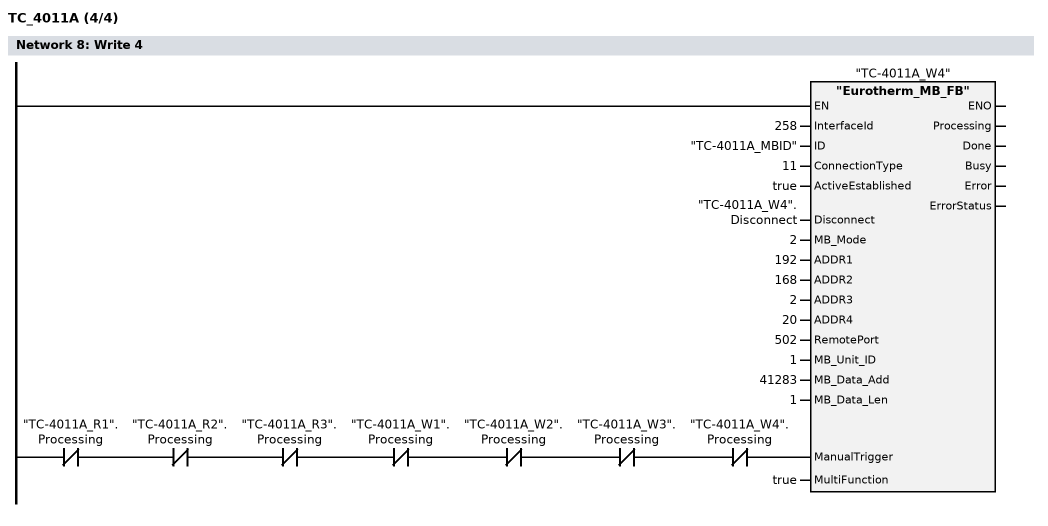
   RUNG wire#powerrail
      "TC-4011A_W4"(ManualTrigger := wire#w1, InterfaceId := 258, ID := "TC-4011A_MBID", ConnectionType := 11, ActiveEstablished := true, Disconnect := "TC-4011A_W4".Disconnect, MB_Mode := 2, ADDR1 := 192, ADDR2 := 168, ADDR3 := 2, ADDR4 := 20, RemotePort := 502, MB_Unit_ID := 1, MB_Data_Add := 41283, MB_Data_Len := 1, MultiFunction := true, Processing =>, Done =>, Busy =>, Error =>, ErrorStatus =>)
   END_RUNG
   RUNG wire#powerrail
      I_Contact( "TC-4011A_R1".Processing )
      I_Contact( "TC-4011A_R2".Processing )
      I_Contact( "TC-4011A_R3".Processing )
      I_Contact( "TC-4011A_W1".Processing )
      I_Contact( "TC-4011A_W2".Processing )
      I_Contact( "TC-4011A_W3".Processing )
      I_Contact( "TC-4011A_W4".Processing )
   END_RUNG wire#w1
   // the same network as SCL:
   "TC-4011A_W4"(InterfaceId := 258,   // "Eurotherm_MB_FB"
                 ID := "TC-4011A_MBID",
                 ConnectionType := 11,
                 ActiveEstablished := true,
                 Disconnect := "TC-4011A_W4".Disconnect,
                 MB_Mode := 2,
                 ADDR1 := 192,
                 ADDR2 := 168,
                 ADDR3 := 2,
                 ADDR4 := 20,
                 RemotePort := 502,
                 MB_Unit_ID := 1,
                 MB_Data_Add := 41283,
                 MB_Data_Len := 1,
                 ManualTrigger := NOT "TC-4011A_R1".Processing AND NOT "TC-4011A_R2".Processing AND NOT "TC-4011A_R3".Processing AND NOT "TC-4011A_W1".Processing AND NOT "TC-4011A_W2".Processing AND NOT "TC-4011A_W3".Processing AND NOT "TC-4011A_W4".Processing,
                 MultiFunction := true);
END_REGION
END_FUNCTION

// folder: Outside Comms/ModBus Comms/EurothermControllers/TC-4011B

FUNCTION "TC_4011B" : Void   // FC32, LAD
{ S7_Optimized_Access := 'TRUE' }
VERSION : 0.1
BEGIN

REGION Network 2: Read Data 1
   // R1=30001
   // R2=31280
   // R3=30023
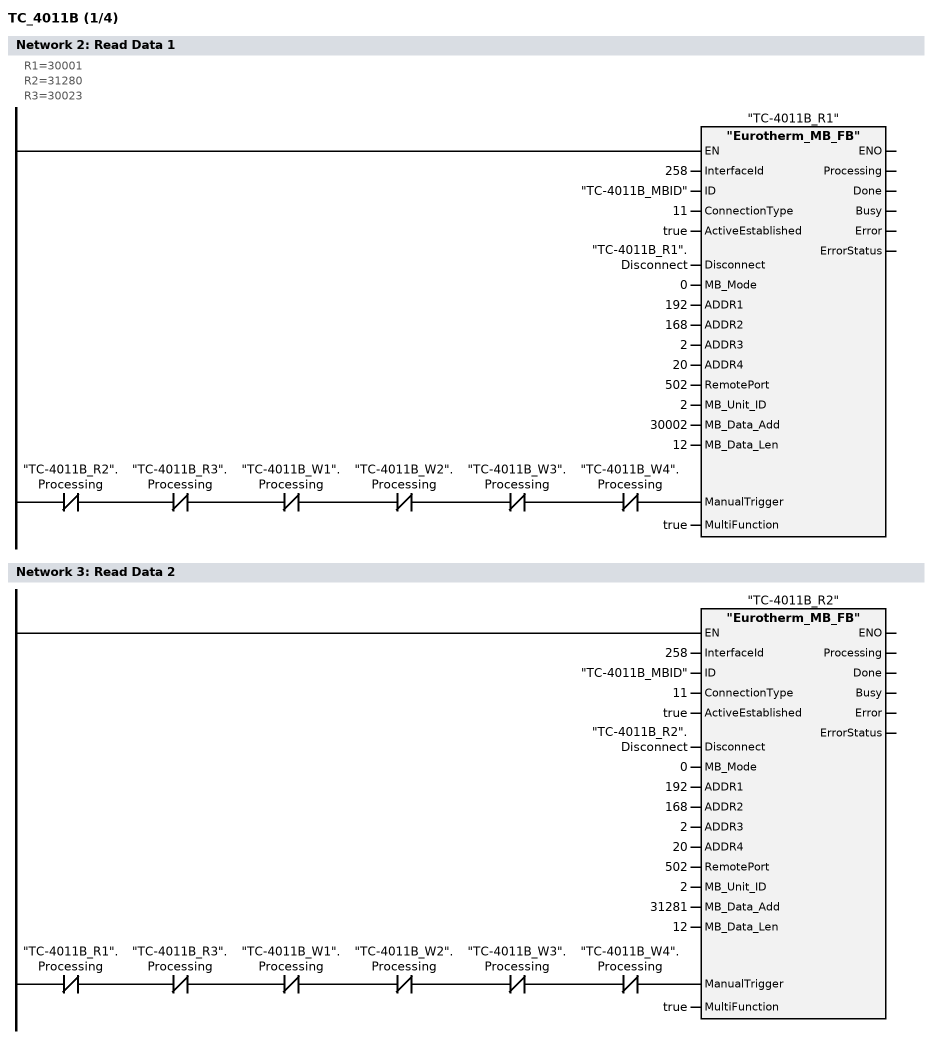
   RUNG wire#powerrail
      "TC-4011B_R1"(ManualTrigger := wire#w1, InterfaceId := 258, ID := "TC-4011B_MBID", ConnectionType := 11, ActiveEstablished := true, Disconnect := "TC-4011B_R1".Disconnect, MB_Mode := 0, ADDR1 := 192, ADDR2 := 168, ADDR3 := 2, ADDR4 := 20, RemotePort := 502, MB_Unit_ID := 2, MB_Data_Add := 30002, MB_Data_Len := 12, MultiFunction := true, Processing =>, Done =>, Busy =>, Error =>, ErrorStatus =>)
   END_RUNG
   RUNG wire#powerrail
      I_Contact( "TC-4011B_R2".Processing )
      I_Contact( "TC-4011B_R3".Processing )
      I_Contact( "TC-4011B_W1".Processing )
      I_Contact( "TC-4011B_W2".Processing )
      I_Contact( "TC-4011B_W3".Processing )
      I_Contact( "TC-4011B_W4".Processing )
   END_RUNG wire#w1
   // the same network as SCL:
   "TC-4011B_R1"(InterfaceId := 258,   // "Eurotherm_MB_FB"
                 ID := "TC-4011B_MBID",
                 ConnectionType := 11,
                 ActiveEstablished := true,
                 Disconnect := "TC-4011B_R1".Disconnect,
                 MB_Mode := 0,
                 ADDR1 := 192,
                 ADDR2 := 168,
                 ADDR3 := 2,
                 ADDR4 := 20,
                 RemotePort := 502,
                 MB_Unit_ID := 2,
                 MB_Data_Add := 30002,
                 MB_Data_Len := 12,
                 ManualTrigger := NOT "TC-4011B_R2".Processing AND NOT "TC-4011B_R3".Processing AND NOT "TC-4011B_W1".Processing AND NOT "TC-4011B_W2".Processing AND NOT "TC-4011B_W3".Processing AND NOT "TC-4011B_W4".Processing,
                 MultiFunction := true);
END_REGION

REGION Network 3: Read Data 2
   RUNG wire#powerrail
      "TC-4011B_R2"(ManualTrigger := wire#w1, InterfaceId := 258, ID := "TC-4011B_MBID", ConnectionType := 11, ActiveEstablished := true, Disconnect := "TC-4011B_R2".Disconnect, MB_Mode := 0, ADDR1 := 192, ADDR2 := 168, ADDR3 := 2, ADDR4 := 20, RemotePort := 502, MB_Unit_ID := 2, MB_Data_Add := 31281, MB_Data_Len := 12, MultiFunction := true, Processing =>, Done =>, Busy =>, Error =>, ErrorStatus =>)
   END_RUNG
   RUNG wire#powerrail
      I_Contact( "TC-4011B_R1".Processing )
      I_Contact( "TC-4011B_R3".Processing )
      I_Contact( "TC-4011B_W1".Processing )
      I_Contact( "TC-4011B_W2".Processing )
      I_Contact( "TC-4011B_W3".Processing )
      I_Contact( "TC-4011B_W4".Processing )
   END_RUNG wire#w1
   // the same network as SCL:
   "TC-4011B_R2"(InterfaceId := 258,   // "Eurotherm_MB_FB"
                 ID := "TC-4011B_MBID",
                 ConnectionType := 11,
                 ActiveEstablished := true,
                 Disconnect := "TC-4011B_R2".Disconnect,
                 MB_Mode := 0,
                 ADDR1 := 192,
                 ADDR2 := 168,
                 ADDR3 := 2,
                 ADDR4 := 20,
                 RemotePort := 502,
                 MB_Unit_ID := 2,
                 MB_Data_Add := 31281,
                 MB_Data_Len := 12,
                 ManualTrigger := NOT "TC-4011B_R1".Processing AND NOT "TC-4011B_R3".Processing AND NOT "TC-4011B_W1".Processing AND NOT "TC-4011B_W2".Processing AND NOT "TC-4011B_W3".Processing AND NOT "TC-4011B_W4".Processing,
                 MultiFunction := true);
END_REGION

REGION Network 4: Read Data 3
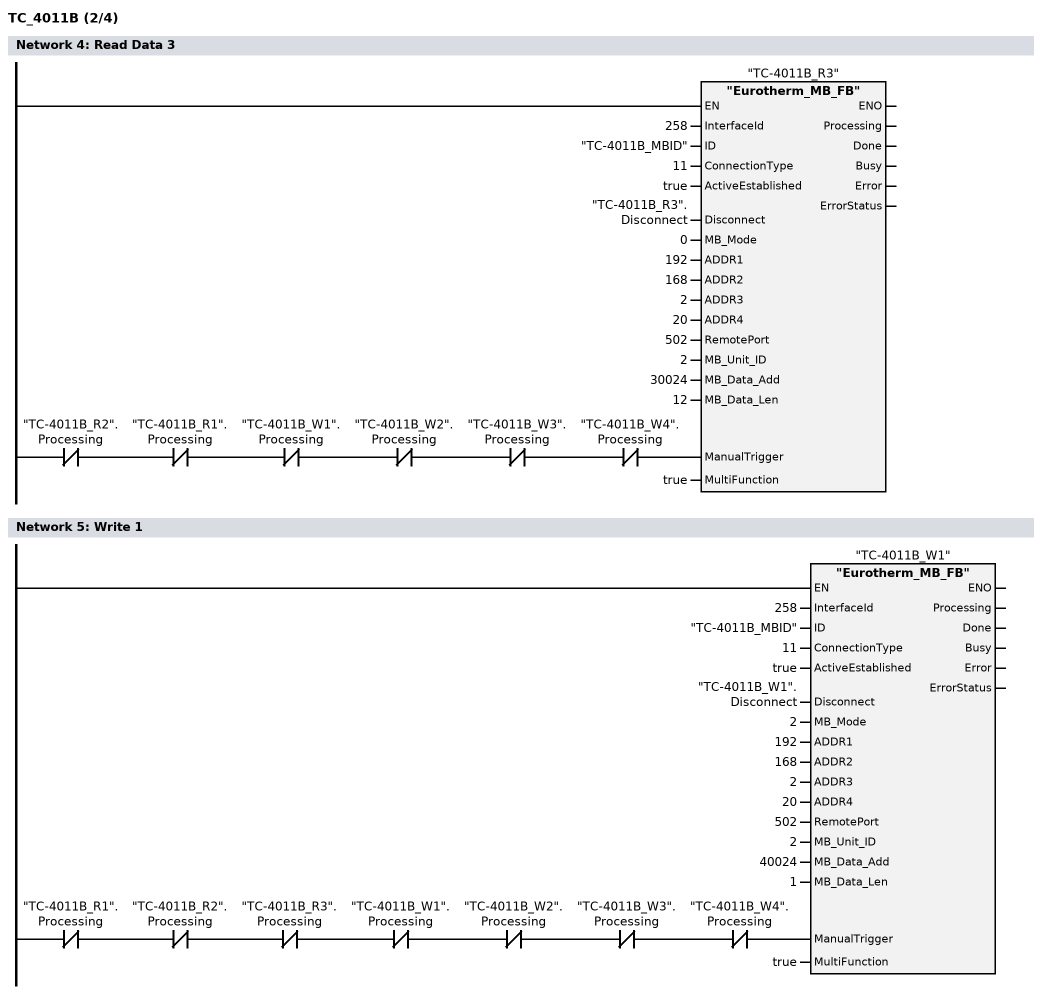
   RUNG wire#powerrail
      "TC-4011B_R3"(ManualTrigger := wire#w1, InterfaceId := 258, ID := "TC-4011B_MBID", ConnectionType := 11, ActiveEstablished := true, Disconnect := "TC-4011B_R3".Disconnect, MB_Mode := 0, ADDR1 := 192, ADDR2 := 168, ADDR3 := 2, ADDR4 := 20, RemotePort := 502, MB_Unit_ID := 2, MB_Data_Add := 30024, MB_Data_Len := 12, MultiFunction := true, Processing =>, Done =>, Busy =>, Error =>, ErrorStatus =>)
   END_RUNG
   RUNG wire#powerrail
      I_Contact( "TC-4011B_R2".Processing )
      I_Contact( "TC-4011B_R1".Processing )
      I_Contact( "TC-4011B_W1".Processing )
      I_Contact( "TC-4011B_W2".Processing )
      I_Contact( "TC-4011B_W3".Processing )
      I_Contact( "TC-4011B_W4".Processing )
   END_RUNG wire#w1
   // the same network as SCL:
   "TC-4011B_R3"(InterfaceId := 258,   // "Eurotherm_MB_FB"
                 ID := "TC-4011B_MBID",
                 ConnectionType := 11,
                 ActiveEstablished := true,
                 Disconnect := "TC-4011B_R3".Disconnect,
                 MB_Mode := 0,
                 ADDR1 := 192,
                 ADDR2 := 168,
                 ADDR3 := 2,
                 ADDR4 := 20,
                 RemotePort := 502,
                 MB_Unit_ID := 2,
                 MB_Data_Add := 30024,
                 MB_Data_Len := 12,
                 ManualTrigger := NOT "TC-4011B_R2".Processing AND NOT "TC-4011B_R1".Processing AND NOT "TC-4011B_W1".Processing AND NOT "TC-4011B_W2".Processing AND NOT "TC-4011B_W3".Processing AND NOT "TC-4011B_W4".Processing,
                 MultiFunction := true);
END_REGION

REGION Network 5: Write 1
   RUNG wire#powerrail
      "TC-4011B_W1"(ManualTrigger := wire#w1, InterfaceId := 258, ID := "TC-4011B_MBID", ConnectionType := 11, ActiveEstablished := true, Disconnect := "TC-4011B_W1".Disconnect, MB_Mode := 2, ADDR1 := 192, ADDR2 := 168, ADDR3 := 2, ADDR4 := 20, RemotePort := 502, MB_Unit_ID := 2, MB_Data_Add := 40024, MB_Data_Len := 1, MultiFunction := true, Processing =>, Done =>, Busy =>, Error =>, ErrorStatus =>)
   END_RUNG
   RUNG wire#powerrail
      I_Contact( "TC-4011B_R1".Processing )
      I_Contact( "TC-4011B_R2".Processing )
      I_Contact( "TC-4011B_R3".Processing )
      I_Contact( "TC-4011B_W1".Processing )
      I_Contact( "TC-4011B_W2".Processing )
      I_Contact( "TC-4011B_W3".Processing )
      I_Contact( "TC-4011B_W4".Processing )
   END_RUNG wire#w1
   // the same network as SCL:
   "TC-4011B_W1"(InterfaceId := 258,   // "Eurotherm_MB_FB"
                 ID := "TC-4011B_MBID",
                 ConnectionType := 11,
                 ActiveEstablished := true,
                 Disconnect := "TC-4011B_W1".Disconnect,
                 MB_Mode := 2,
                 ADDR1 := 192,
                 ADDR2 := 168,
                 ADDR3 := 2,
                 ADDR4 := 20,
                 RemotePort := 502,
                 MB_Unit_ID := 2,
                 MB_Data_Add := 40024,
                 MB_Data_Len := 1,
                 ManualTrigger := NOT "TC-4011B_R1".Processing AND NOT "TC-4011B_R2".Processing AND NOT "TC-4011B_R3".Processing AND NOT "TC-4011B_W1".Processing AND NOT "TC-4011B_W2".Processing AND NOT "TC-4011B_W3".Processing AND NOT "TC-4011B_W4".Processing,
                 MultiFunction := true);
END_REGION

REGION Network 6: Write 2
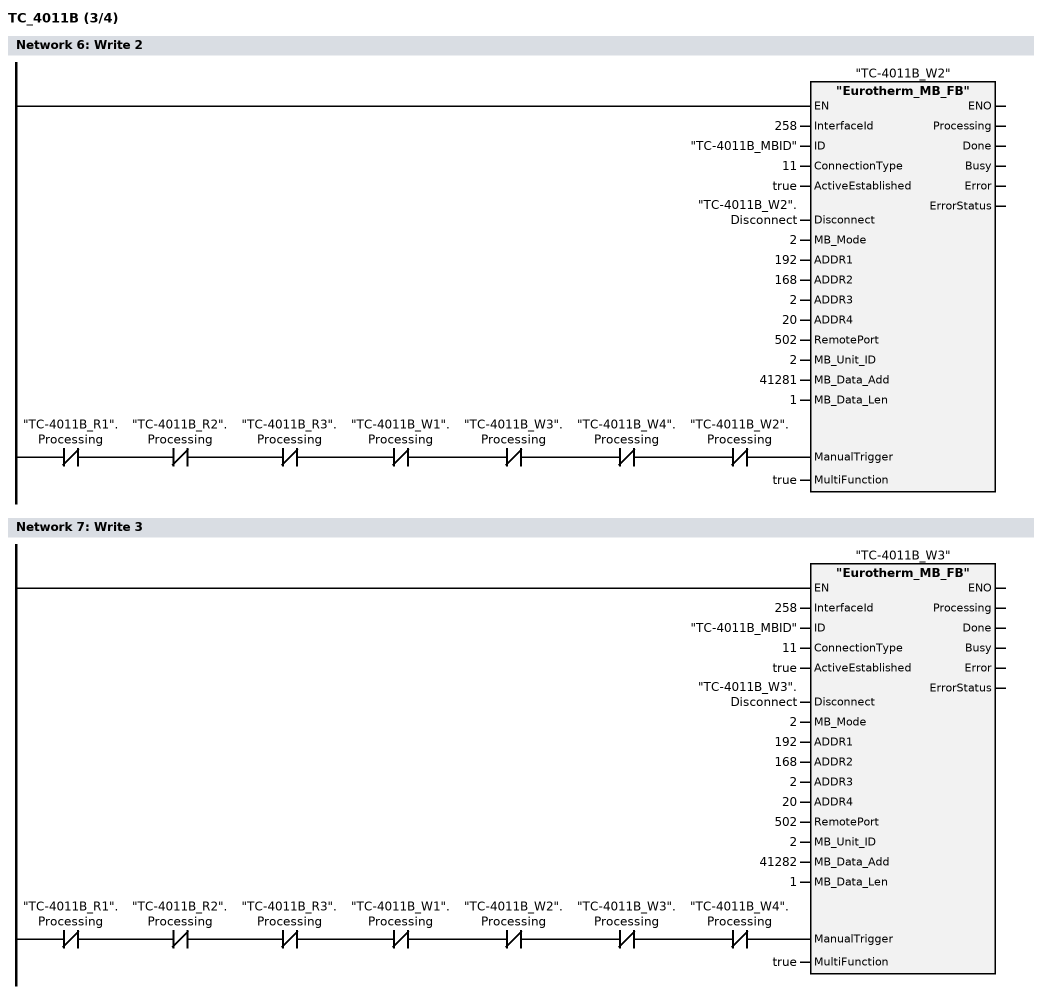
   RUNG wire#powerrail
      "TC-4011B_W2"(ManualTrigger := wire#w1, InterfaceId := 258, ID := "TC-4011B_MBID", ConnectionType := 11, ActiveEstablished := true, Disconnect := "TC-4011B_W2".Disconnect, MB_Mode := 2, ADDR1 := 192, ADDR2 := 168, ADDR3 := 2, ADDR4 := 20, RemotePort := 502, MB_Unit_ID := 2, MB_Data_Add := 41281, MB_Data_Len := 1, MultiFunction := true, Processing =>, Done =>, Busy =>, Error =>, ErrorStatus =>)
   END_RUNG
   RUNG wire#powerrail
      I_Contact( "TC-4011B_R1".Processing )
      I_Contact( "TC-4011B_R2".Processing )
      I_Contact( "TC-4011B_R3".Processing )
      I_Contact( "TC-4011B_W1".Processing )
      I_Contact( "TC-4011B_W3".Processing )
      I_Contact( "TC-4011B_W4".Processing )
      I_Contact( "TC-4011B_W2".Processing )
   END_RUNG wire#w1
   // the same network as SCL:
   "TC-4011B_W2"(InterfaceId := 258,   // "Eurotherm_MB_FB"
                 ID := "TC-4011B_MBID",
                 ConnectionType := 11,
                 ActiveEstablished := true,
                 Disconnect := "TC-4011B_W2".Disconnect,
                 MB_Mode := 2,
                 ADDR1 := 192,
                 ADDR2 := 168,
                 ADDR3 := 2,
                 ADDR4 := 20,
                 RemotePort := 502,
                 MB_Unit_ID := 2,
                 MB_Data_Add := 41281,
                 MB_Data_Len := 1,
                 ManualTrigger := NOT "TC-4011B_R1".Processing AND NOT "TC-4011B_R2".Processing AND NOT "TC-4011B_R3".Processing AND NOT "TC-4011B_W1".Processing AND NOT "TC-4011B_W3".Processing AND NOT "TC-4011B_W4".Processing AND NOT "TC-4011B_W2".Processing,
                 MultiFunction := true);
END_REGION

REGION Network 7: Write 3
   RUNG wire#powerrail
      "TC-4011B_W3"(ManualTrigger := wire#w1, InterfaceId := 258, ID := "TC-4011B_MBID", ConnectionType := 11, ActiveEstablished := true, Disconnect := "TC-4011B_W3".Disconnect, MB_Mode := 2, ADDR1 := 192, ADDR2 := 168, ADDR3 := 2, ADDR4 := 20, RemotePort := 502, MB_Unit_ID := 2, MB_Data_Add := 41282, MB_Data_Len := 1, MultiFunction := true, Processing =>, Done =>, Busy =>, Error =>, ErrorStatus =>)
   END_RUNG
   RUNG wire#powerrail
      I_Contact( "TC-4011B_R1".Processing )
      I_Contact( "TC-4011B_R2".Processing )
      I_Contact( "TC-4011B_R3".Processing )
      I_Contact( "TC-4011B_W1".Processing )
      I_Contact( "TC-4011B_W2".Processing )
      I_Contact( "TC-4011B_W3".Processing )
      I_Contact( "TC-4011B_W4".Processing )
   END_RUNG wire#w1
   // the same network as SCL:
   "TC-4011B_W3"(InterfaceId := 258,   // "Eurotherm_MB_FB"
                 ID := "TC-4011B_MBID",
                 ConnectionType := 11,
                 ActiveEstablished := true,
                 Disconnect := "TC-4011B_W3".Disconnect,
                 MB_Mode := 2,
                 ADDR1 := 192,
                 ADDR2 := 168,
                 ADDR3 := 2,
                 ADDR4 := 20,
                 RemotePort := 502,
                 MB_Unit_ID := 2,
                 MB_Data_Add := 41282,
                 MB_Data_Len := 1,
                 ManualTrigger := NOT "TC-4011B_R1".Processing AND NOT "TC-4011B_R2".Processing AND NOT "TC-4011B_R3".Processing AND NOT "TC-4011B_W1".Processing AND NOT "TC-4011B_W2".Processing AND NOT "TC-4011B_W3".Processing AND NOT "TC-4011B_W4".Processing,
                 MultiFunction := true);
END_REGION

REGION Network 8: Write 4
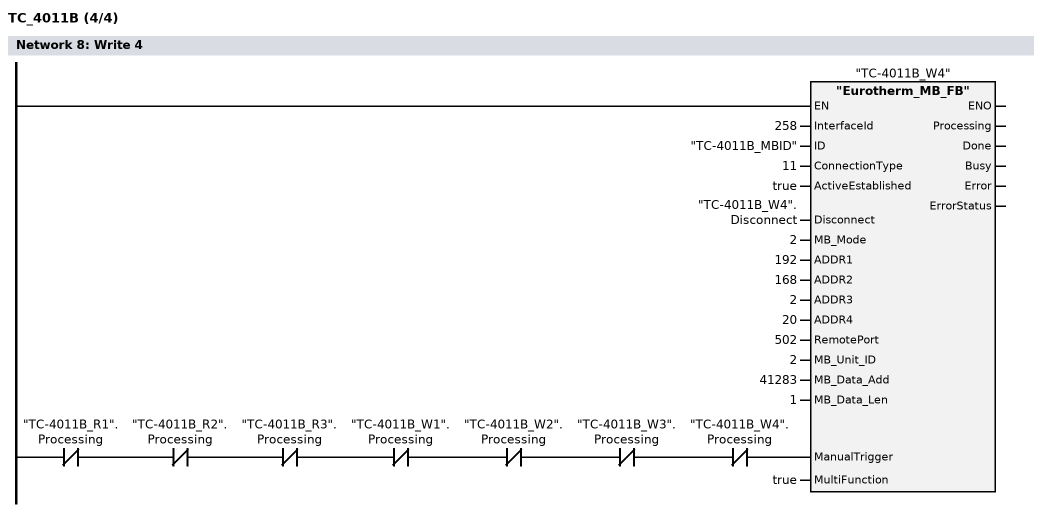
   RUNG wire#powerrail
      "TC-4011B_W4"(ManualTrigger := wire#w1, InterfaceId := 258, ID := "TC-4011B_MBID", ConnectionType := 11, ActiveEstablished := true, Disconnect := "TC-4011B_W4".Disconnect, MB_Mode := 2, ADDR1 := 192, ADDR2 := 168, ADDR3 := 2, ADDR4 := 20, RemotePort := 502, MB_Unit_ID := 2, MB_Data_Add := 41283, MB_Data_Len := 1, MultiFunction := true, Processing =>, Done =>, Busy =>, Error =>, ErrorStatus =>)
   END_RUNG
   RUNG wire#powerrail
      I_Contact( "TC-4011B_R1".Processing )
      I_Contact( "TC-4011B_R2".Processing )
      I_Contact( "TC-4011B_R3".Processing )
      I_Contact( "TC-4011B_W1".Processing )
      I_Contact( "TC-4011B_W2".Processing )
      I_Contact( "TC-4011B_W3".Processing )
      I_Contact( "TC-4011B_W4".Processing )
   END_RUNG wire#w1
   // the same network as SCL:
   "TC-4011B_W4"(InterfaceId := 258,   // "Eurotherm_MB_FB"
                 ID := "TC-4011B_MBID",
                 ConnectionType := 11,
                 ActiveEstablished := true,
                 Disconnect := "TC-4011B_W4".Disconnect,
                 MB_Mode := 2,
                 ADDR1 := 192,
                 ADDR2 := 168,
                 ADDR3 := 2,
                 ADDR4 := 20,
                 RemotePort := 502,
                 MB_Unit_ID := 2,
                 MB_Data_Add := 41283,
                 MB_Data_Len := 1,
                 ManualTrigger := NOT "TC-4011B_R1".Processing AND NOT "TC-4011B_R2".Processing AND NOT "TC-4011B_R3".Processing AND NOT "TC-4011B_W1".Processing AND NOT "TC-4011B_W2".Processing AND NOT "TC-4011B_W3".Processing AND NOT "TC-4011B_W4".Processing,
                 MultiFunction := true);
END_REGION
END_FUNCTION

// folder: Outside Comms/ModBus Comms/EurothermControllers/TC-4011C

FUNCTION "TC_4011C" : Void   // FC33, LAD
{ S7_Optimized_Access := 'TRUE' }
VERSION : 0.1
BEGIN

REGION Network 2: Read Data 1
   // R1=30001
   // R2=31280
   // R3=30023
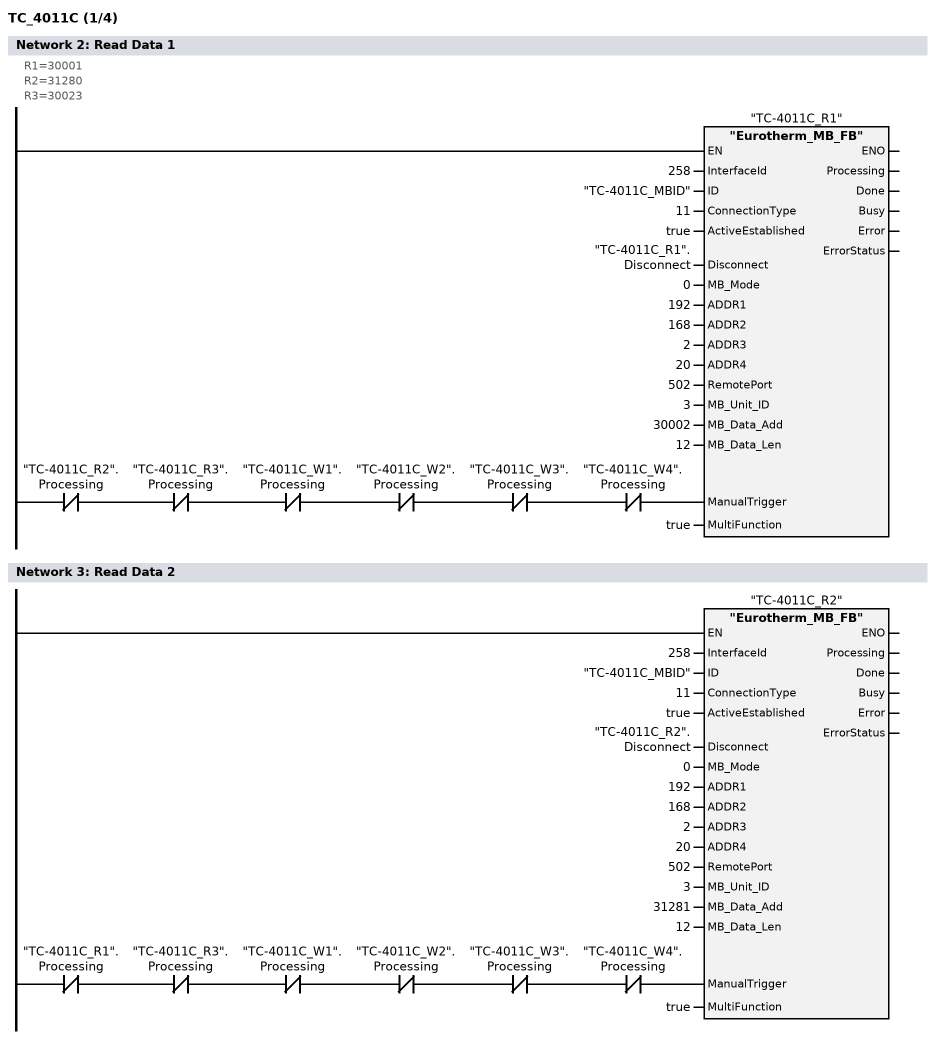
   RUNG wire#powerrail
      "TC-4011C_R1"(ManualTrigger := wire#w1, InterfaceId := 258, ID := "TC-4011C_MBID", ConnectionType := 11, ActiveEstablished := true, Disconnect := "TC-4011C_R1".Disconnect, MB_Mode := 0, ADDR1 := 192, ADDR2 := 168, ADDR3 := 2, ADDR4 := 20, RemotePort := 502, MB_Unit_ID := 3, MB_Data_Add := 30002, MB_Data_Len := 12, MultiFunction := true, Processing =>, Done =>, Busy =>, Error =>, ErrorStatus =>)
   END_RUNG
   RUNG wire#powerrail
      I_Contact( "TC-4011C_R2".Processing )
      I_Contact( "TC-4011C_R3".Processing )
      I_Contact( "TC-4011C_W1".Processing )
      I_Contact( "TC-4011C_W2".Processing )
      I_Contact( "TC-4011C_W3".Processing )
      I_Contact( "TC-4011C_W4".Processing )
   END_RUNG wire#w1
   // the same network as SCL:
   "TC-4011C_R1"(InterfaceId := 258,   // "Eurotherm_MB_FB"
                 ID := "TC-4011C_MBID",
                 ConnectionType := 11,
                 ActiveEstablished := true,
                 Disconnect := "TC-4011C_R1".Disconnect,
                 MB_Mode := 0,
                 ADDR1 := 192,
                 ADDR2 := 168,
                 ADDR3 := 2,
                 ADDR4 := 20,
                 RemotePort := 502,
                 MB_Unit_ID := 3,
                 MB_Data_Add := 30002,
                 MB_Data_Len := 12,
                 ManualTrigger := NOT "TC-4011C_R2".Processing AND NOT "TC-4011C_R3".Processing AND NOT "TC-4011C_W1".Processing AND NOT "TC-4011C_W2".Processing AND NOT "TC-4011C_W3".Processing AND NOT "TC-4011C_W4".Processing,
                 MultiFunction := true);
END_REGION

REGION Network 3: Read Data 2
   RUNG wire#powerrail
      "TC-4011C_R2"(ManualTrigger := wire#w1, InterfaceId := 258, ID := "TC-4011C_MBID", ConnectionType := 11, ActiveEstablished := true, Disconnect := "TC-4011C_R2".Disconnect, MB_Mode := 0, ADDR1 := 192, ADDR2 := 168, ADDR3 := 2, ADDR4 := 20, RemotePort := 502, MB_Unit_ID := 3, MB_Data_Add := 31281, MB_Data_Len := 12, MultiFunction := true, Processing =>, Done =>, Busy =>, Error =>, ErrorStatus =>)
   END_RUNG
   RUNG wire#powerrail
      I_Contact( "TC-4011C_R1".Processing )
      I_Contact( "TC-4011C_R3".Processing )
      I_Contact( "TC-4011C_W1".Processing )
      I_Contact( "TC-4011C_W2".Processing )
      I_Contact( "TC-4011C_W3".Processing )
      I_Contact( "TC-4011C_W4".Processing )
   END_RUNG wire#w1
   // the same network as SCL:
   "TC-4011C_R2"(InterfaceId := 258,   // "Eurotherm_MB_FB"
                 ID := "TC-4011C_MBID",
                 ConnectionType := 11,
                 ActiveEstablished := true,
                 Disconnect := "TC-4011C_R2".Disconnect,
                 MB_Mode := 0,
                 ADDR1 := 192,
                 ADDR2 := 168,
                 ADDR3 := 2,
                 ADDR4 := 20,
                 RemotePort := 502,
                 MB_Unit_ID := 3,
                 MB_Data_Add := 31281,
                 MB_Data_Len := 12,
                 ManualTrigger := NOT "TC-4011C_R1".Processing AND NOT "TC-4011C_R3".Processing AND NOT "TC-4011C_W1".Processing AND NOT "TC-4011C_W2".Processing AND NOT "TC-4011C_W3".Processing AND NOT "TC-4011C_W4".Processing,
                 MultiFunction := true);
END_REGION

REGION Network 4: Read Data 3
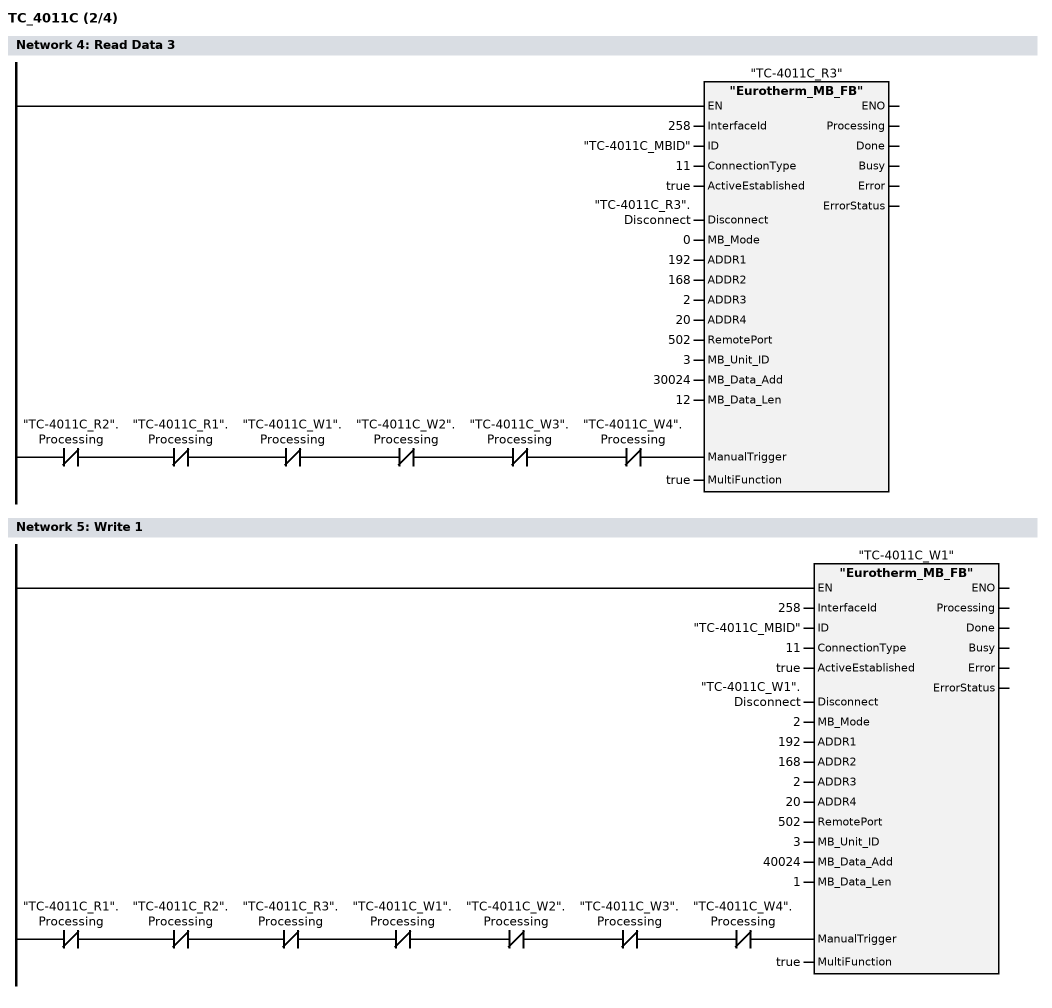
   RUNG wire#powerrail
      "TC-4011C_R3"(ManualTrigger := wire#w1, InterfaceId := 258, ID := "TC-4011C_MBID", ConnectionType := 11, ActiveEstablished := true, Disconnect := "TC-4011C_R3".Disconnect, MB_Mode := 0, ADDR1 := 192, ADDR2 := 168, ADDR3 := 2, ADDR4 := 20, RemotePort := 502, MB_Unit_ID := 3, MB_Data_Add := 30024, MB_Data_Len := 12, MultiFunction := true, Processing =>, Done =>, Busy =>, Error =>, ErrorStatus =>)
   END_RUNG
   RUNG wire#powerrail
      I_Contact( "TC-4011C_R2".Processing )
      I_Contact( "TC-4011C_R1".Processing )
      I_Contact( "TC-4011C_W1".Processing )
      I_Contact( "TC-4011C_W2".Processing )
      I_Contact( "TC-4011C_W3".Processing )
      I_Contact( "TC-4011C_W4".Processing )
   END_RUNG wire#w1
   // the same network as SCL:
   "TC-4011C_R3"(InterfaceId := 258,   // "Eurotherm_MB_FB"
                 ID := "TC-4011C_MBID",
                 ConnectionType := 11,
                 ActiveEstablished := true,
                 Disconnect := "TC-4011C_R3".Disconnect,
                 MB_Mode := 0,
                 ADDR1 := 192,
                 ADDR2 := 168,
                 ADDR3 := 2,
                 ADDR4 := 20,
                 RemotePort := 502,
                 MB_Unit_ID := 3,
                 MB_Data_Add := 30024,
                 MB_Data_Len := 12,
                 ManualTrigger := NOT "TC-4011C_R2".Processing AND NOT "TC-4011C_R1".Processing AND NOT "TC-4011C_W1".Processing AND NOT "TC-4011C_W2".Processing AND NOT "TC-4011C_W3".Processing AND NOT "TC-4011C_W4".Processing,
                 MultiFunction := true);
END_REGION

REGION Network 5: Write 1
   RUNG wire#powerrail
      "TC-4011C_W1"(ManualTrigger := wire#w1, InterfaceId := 258, ID := "TC-4011C_MBID", ConnectionType := 11, ActiveEstablished := true, Disconnect := "TC-4011C_W1".Disconnect, MB_Mode := 2, ADDR1 := 192, ADDR2 := 168, ADDR3 := 2, ADDR4 := 20, RemotePort := 502, MB_Unit_ID := 3, MB_Data_Add := 40024, MB_Data_Len := 1, MultiFunction := true, Processing =>, Done =>, Busy =>, Error =>, ErrorStatus =>)
   END_RUNG
   RUNG wire#powerrail
      I_Contact( "TC-4011C_R1".Processing )
      I_Contact( "TC-4011C_R2".Processing )
      I_Contact( "TC-4011C_R3".Processing )
      I_Contact( "TC-4011C_W1".Processing )
      I_Contact( "TC-4011C_W2".Processing )
      I_Contact( "TC-4011C_W3".Processing )
      I_Contact( "TC-4011C_W4".Processing )
   END_RUNG wire#w1
   // the same network as SCL:
   "TC-4011C_W1"(InterfaceId := 258,   // "Eurotherm_MB_FB"
                 ID := "TC-4011C_MBID",
                 ConnectionType := 11,
                 ActiveEstablished := true,
                 Disconnect := "TC-4011C_W1".Disconnect,
                 MB_Mode := 2,
                 ADDR1 := 192,
                 ADDR2 := 168,
                 ADDR3 := 2,
                 ADDR4 := 20,
                 RemotePort := 502,
                 MB_Unit_ID := 3,
                 MB_Data_Add := 40024,
                 MB_Data_Len := 1,
                 ManualTrigger := NOT "TC-4011C_R1".Processing AND NOT "TC-4011C_R2".Processing AND NOT "TC-4011C_R3".Processing AND NOT "TC-4011C_W1".Processing AND NOT "TC-4011C_W2".Processing AND NOT "TC-4011C_W3".Processing AND NOT "TC-4011C_W4".Processing,
                 MultiFunction := true);
END_REGION

REGION Network 6: Write 2
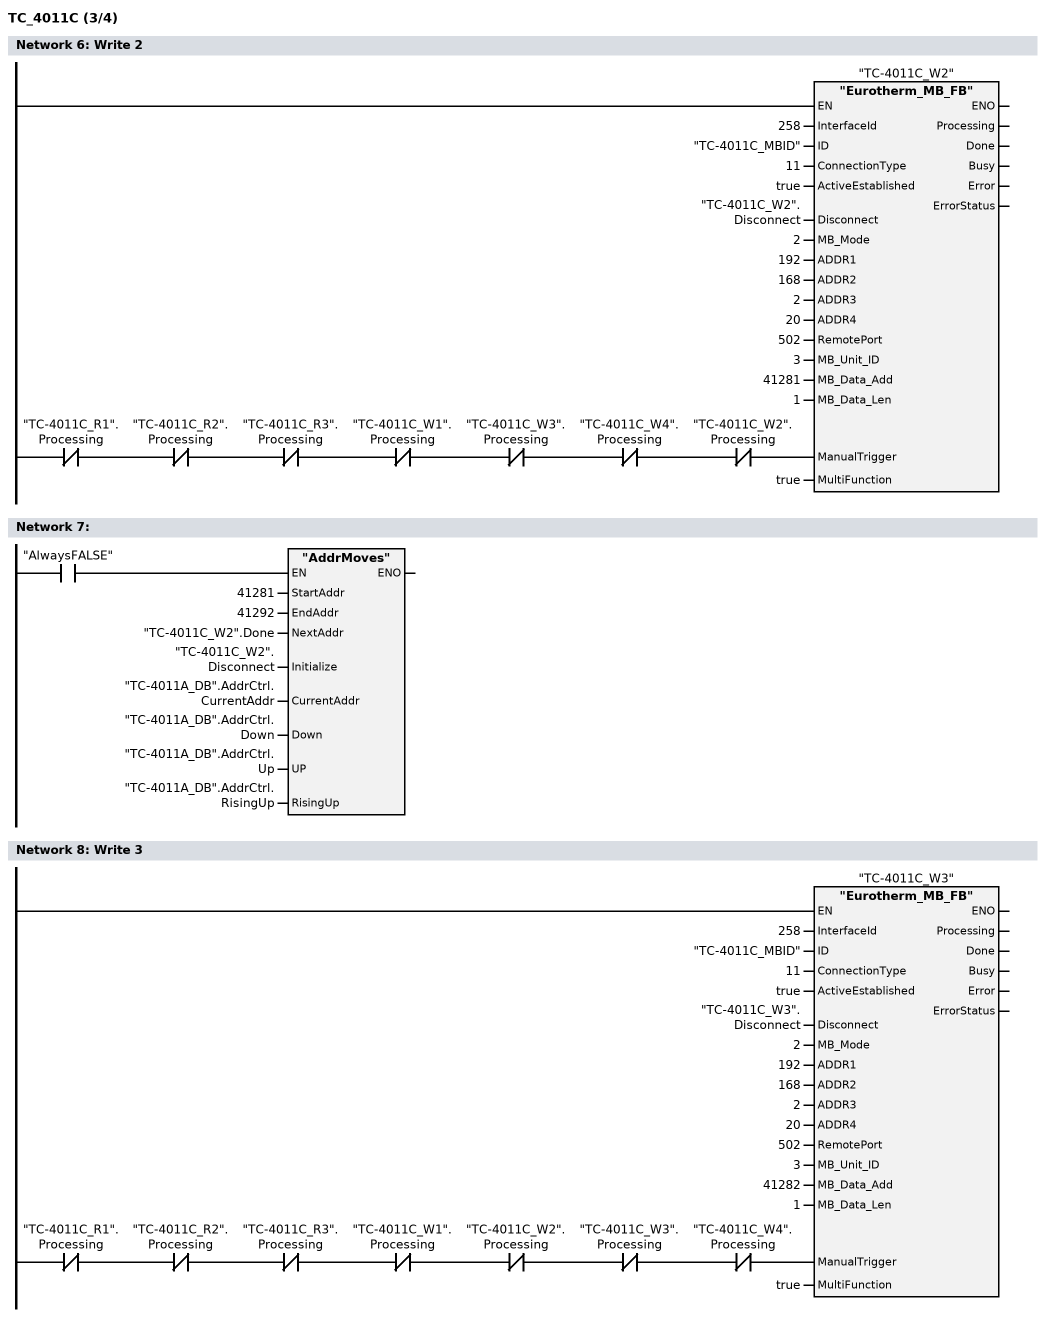
   RUNG wire#powerrail
      "TC-4011C_W2"(ManualTrigger := wire#w1, InterfaceId := 258, ID := "TC-4011C_MBID", ConnectionType := 11, ActiveEstablished := true, Disconnect := "TC-4011C_W2".Disconnect, MB_Mode := 2, ADDR1 := 192, ADDR2 := 168, ADDR3 := 2, ADDR4 := 20, RemotePort := 502, MB_Unit_ID := 3, MB_Data_Add := 41281, MB_Data_Len := 1, MultiFunction := true, Processing =>, Done =>, Busy =>, Error =>, ErrorStatus =>)
   END_RUNG
   RUNG wire#powerrail
      I_Contact( "TC-4011C_R1".Processing )
      I_Contact( "TC-4011C_R2".Processing )
      I_Contact( "TC-4011C_R3".Processing )
      I_Contact( "TC-4011C_W1".Processing )
      I_Contact( "TC-4011C_W3".Processing )
      I_Contact( "TC-4011C_W4".Processing )
      I_Contact( "TC-4011C_W2".Processing )
   END_RUNG wire#w1
   // the same network as SCL:
   "TC-4011C_W2"(InterfaceId := 258,   // "Eurotherm_MB_FB"